// TIA Portal project "FABRICA DE TAPAS - TRANSPORTE -TUNEL DE ENFRIAMIENTO" (V17) (continued)
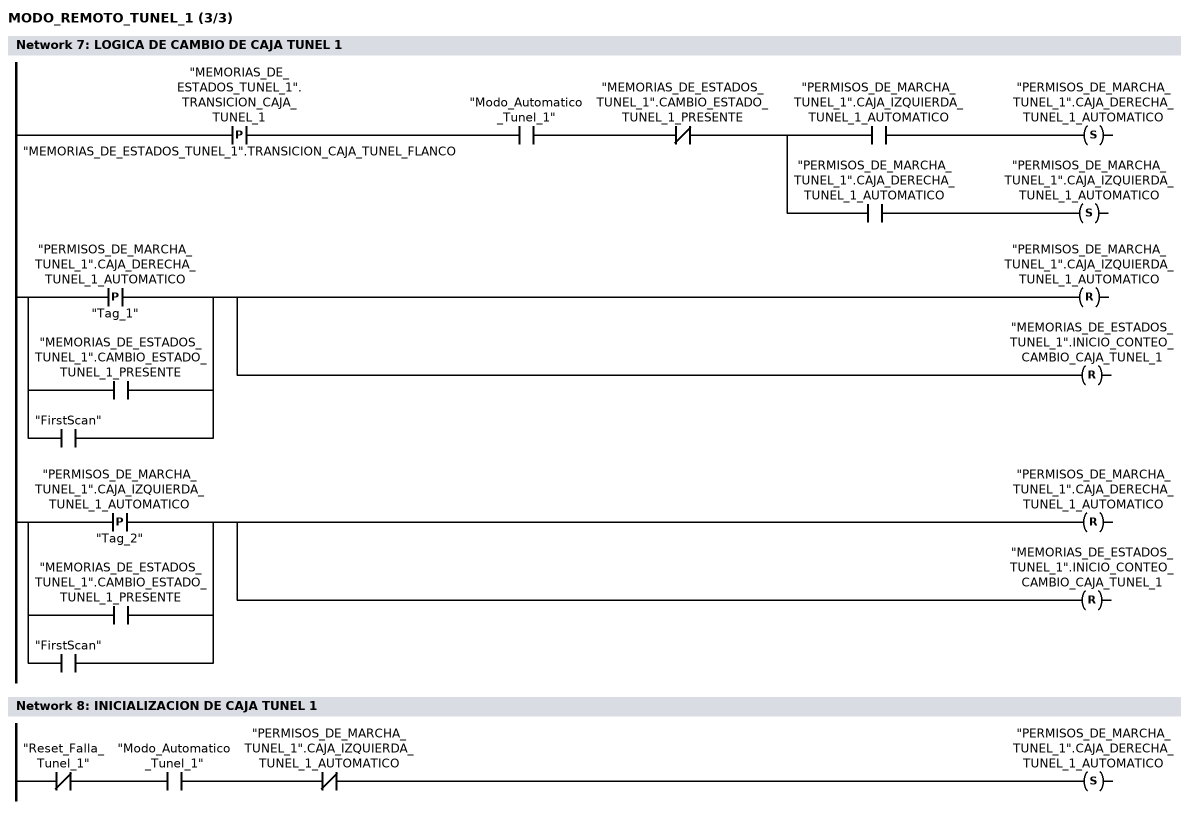
   RUNG wire#powerrail
      P_Contact(operand := "MEMORIAS_DE_ESTADOS_TUNEL_1".TRANSICION_CAJA_TUNEL_1, bit := "MEMORIAS_DE_ESTADOS_TUNEL_1".TRANSICION_CAJA_TUNEL_FLANCO)
      Contact( "Modo_Automatico_Tunel_1" )
      I_Contact( "MEMORIAS_DE_ESTADOS_TUNEL_1".CAMBIO_ESTADO_TUNEL_1_PRESENTE )
      wire#w1
      Contact( "PERMISOS_DE_MARCHA_TUNEL_1".CAJA_IZQUIERDA_TUNEL_1_AUTOMATICO )
      S_Coil( "PERMISOS_DE_MARCHA_TUNEL_1".CAJA_DERECHA_TUNEL_1_AUTOMATICO )
   END_RUNG
   RUNG wire#w1
      Contact( "PERMISOS_DE_MARCHA_TUNEL_1".CAJA_DERECHA_TUNEL_1_AUTOMATICO )
      S_Coil( "PERMISOS_DE_MARCHA_TUNEL_1".CAJA_IZQUIERDA_TUNEL_1_AUTOMATICO )
   END_RUNG
   RUNG wire#powerrail
      P_Contact(operand := "PERMISOS_DE_MARCHA_TUNEL_1".CAJA_DERECHA_TUNEL_1_AUTOMATICO, bit := "Tag_1")
      wire#w2
      R_Coil( "PERMISOS_DE_MARCHA_TUNEL_1".CAJA_IZQUIERDA_TUNEL_1_AUTOMATICO )
   END_RUNG
   RUNG wire#powerrail
      Contact( "MEMORIAS_DE_ESTADOS_TUNEL_1".CAMBIO_ESTADO_TUNEL_1_PRESENTE )
   END_RUNG wire#w2
   RUNG wire#powerrail
      Contact( "FirstScan" )
   END_RUNG wire#w2
   RUNG wire#w2
      R_Coil( "MEMORIAS_DE_ESTADOS_TUNEL_1".INICIO_CONTEO_CAMBIO_CAJA_TUNEL_1 )
   END_RUNG
   RUNG wire#powerrail
      P_Contact(operand := "PERMISOS_DE_MARCHA_TUNEL_1".CAJA_IZQUIERDA_TUNEL_1_AUTOMATICO, bit := "Tag_2")
      wire#w3
      R_Coil( "PERMISOS_DE_MARCHA_TUNEL_1".CAJA_DERECHA_TUNEL_1_AUTOMATICO )
   END_RUNG
   RUNG wire#powerrail
      Contact( "MEMORIAS_DE_ESTADOS_TUNEL_1".CAMBIO_ESTADO_TUNEL_1_PRESENTE )
   END_RUNG wire#w3
   RUNG wire#powerrail
      Contact( "FirstScan" )
   END_RUNG wire#w3
   RUNG wire#w3
      R_Coil( "MEMORIAS_DE_ESTADOS_TUNEL_1".INICIO_CONTEO_CAMBIO_CAJA_TUNEL_1 )
   END_RUNG
   // the same network as SCL:
   #_w1 := "MEMORIAS_DE_ESTADOS_TUNEL_1".TRANSICION_CAJA_TUNEL_1 AND NOT "MEMORIAS_DE_ESTADOS_TUNEL_1".TRANSICION_CAJA_TUNEL_FLANCO;   // rising edge of "MEMORIAS_DE_ESTADOS_TUNEL_1".TRANSICION_CAJA_TUNEL_1
   "MEMORIAS_DE_ESTADOS_TUNEL_1".TRANSICION_CAJA_TUNEL_FLANCO := "MEMORIAS_DE_ESTADOS_TUNEL_1".TRANSICION_CAJA_TUNEL_1;
   #_w2 := #_w1 AND "Modo_Automatico_Tunel_1" AND NOT "MEMORIAS_DE_ESTADOS_TUNEL_1".CAMBIO_ESTADO_TUNEL_1_PRESENTE;
   IF #_w2 AND "PERMISOS_DE_MARCHA_TUNEL_1".CAJA_IZQUIERDA_TUNEL_1_AUTOMATICO THEN
       "PERMISOS_DE_MARCHA_TUNEL_1".CAJA_DERECHA_TUNEL_1_AUTOMATICO := TRUE;
   END_IF;
   IF #_w2 AND "PERMISOS_DE_MARCHA_TUNEL_1".CAJA_DERECHA_TUNEL_1_AUTOMATICO THEN
       "PERMISOS_DE_MARCHA_TUNEL_1".CAJA_IZQUIERDA_TUNEL_1_AUTOMATICO := TRUE;
   END_IF;
   #_w3 := "PERMISOS_DE_MARCHA_TUNEL_1".CAJA_DERECHA_TUNEL_1_AUTOMATICO AND NOT "Tag_1";   // rising edge of "PERMISOS_DE_MARCHA_TUNEL_1".CAJA_DERECHA_TUNEL_1_AUTOMATICO
   "Tag_1" := "PERMISOS_DE_MARCHA_TUNEL_1".CAJA_DERECHA_TUNEL_1_AUTOMATICO;
   IF #_w3 OR "MEMORIAS_DE_ESTADOS_TUNEL_1".CAMBIO_ESTADO_TUNEL_1_PRESENTE OR "FirstScan" THEN
       "PERMISOS_DE_MARCHA_TUNEL_1".CAJA_IZQUIERDA_TUNEL_1_AUTOMATICO := FALSE;
       "MEMORIAS_DE_ESTADOS_TUNEL_1".INICIO_CONTEO_CAMBIO_CAJA_TUNEL_1 := FALSE;
   END_IF;
   #_w4 := "PERMISOS_DE_MARCHA_TUNEL_1".CAJA_IZQUIERDA_TUNEL_1_AUTOMATICO AND NOT "Tag_2";   // rising edge of "PERMISOS_DE_MARCHA_TUNEL_1".CAJA_IZQUIERDA_TUNEL_1_AUTOMATICO
   "Tag_2" := "PERMISOS_DE_MARCHA_TUNEL_1".CAJA_IZQUIERDA_TUNEL_1_AUTOMATICO;
   IF #_w4 OR "MEMORIAS_DE_ESTADOS_TUNEL_1".CAMBIO_ESTADO_TUNEL_1_PRESENTE OR "FirstScan" THEN
       "PERMISOS_DE_MARCHA_TUNEL_1".CAJA_DERECHA_TUNEL_1_AUTOMATICO := FALSE;
       "MEMORIAS_DE_ESTADOS_TUNEL_1".INICIO_CONTEO_CAMBIO_CAJA_TUNEL_1 := FALSE;
   END_IF;
END_REGION

REGION Network 8: INICIALIZACION DE CAJA TUNEL 1
   RUNG wire#powerrail
      I_Contact( "Reset_Falla_Tunel_1" )
      Contact( "Modo_Automatico_Tunel_1" )
      I_Contact( "PERMISOS_DE_MARCHA_TUNEL_1".CAJA_IZQUIERDA_TUNEL_1_AUTOMATICO )
      S_Coil( "PERMISOS_DE_MARCHA_TUNEL_1".CAJA_DERECHA_TUNEL_1_AUTOMATICO )
   END_RUNG
   // the same network as SCL:
   IF NOT "Reset_Falla_Tunel_1" AND "Modo_Automatico_Tunel_1" AND NOT "PERMISOS_DE_MARCHA_TUNEL_1".CAJA_IZQUIERDA_TUNEL_1_AUTOMATICO THEN
       "PERMISOS_DE_MARCHA_TUNEL_1".CAJA_DERECHA_TUNEL_1_AUTOMATICO := TRUE;
   END_IF;
END_REGION
END_FUNCTION

FUNCTION "MODO_REMOTO_TUNEL_2" : Void   // FC2, LAD
{ S7_Optimized_Access := 'TRUE' }
VERSION : 0.1
   VAR_TEMP   // added for the SCL form of the ladder/FBD networks
      _w1 : Bool;
      _w2 : Bool;
      _w3 : Bool;
      _w4 : Bool;
   END_VAR
BEGIN

REGION Network 1
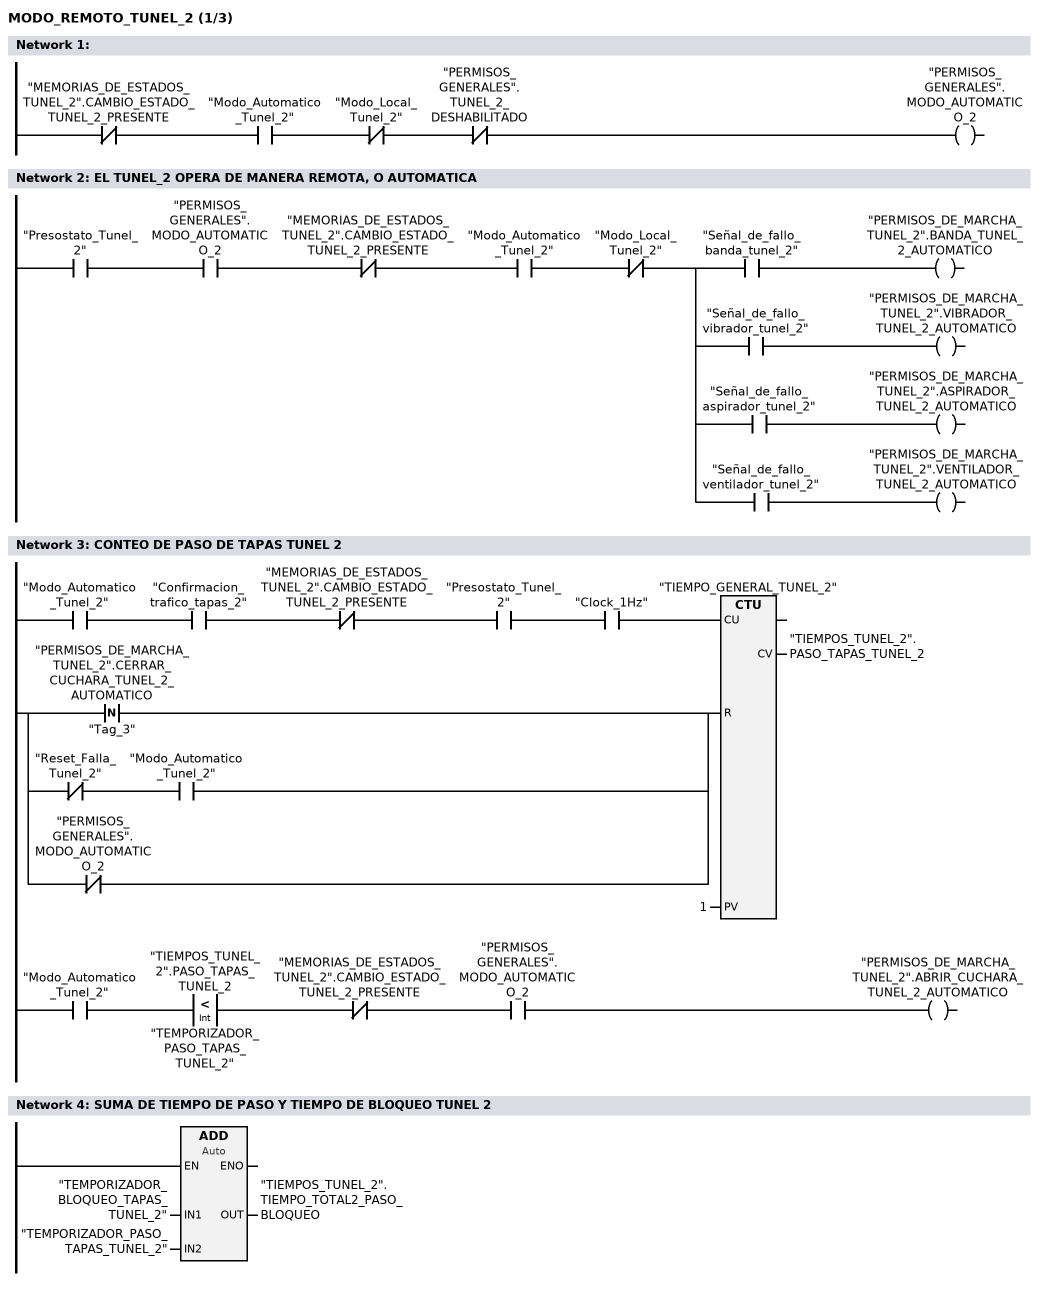
   RUNG wire#powerrail
      I_Contact( "MEMORIAS_DE_ESTADOS_TUNEL_2".CAMBIO_ESTADO_TUNEL_2_PRESENTE )
      Contact( "Modo_Automatico_Tunel_2" )
      I_Contact( "Modo_Local_Tunel_2" )
      I_Contact( "PERMISOS_GENERALES".TUNEL_2_DESHABILITADO )
      Coil( "PERMISOS_GENERALES".MODO_AUTOMATICO_2 )
   END_RUNG
   // the same network as SCL:
   "PERMISOS_GENERALES".MODO_AUTOMATICO_2 := NOT "MEMORIAS_DE_ESTADOS_TUNEL_2".CAMBIO_ESTADO_TUNEL_2_PRESENTE AND "Modo_Automatico_Tunel_2" AND NOT "Modo_Local_Tunel_2" AND NOT "PERMISOS_GENERALES".TUNEL_2_DESHABILITADO;
END_REGION

REGION Network 2: EL TUNEL_2 OPERA DE MANERA REMOTA, O AUTOMATICA
   RUNG wire#powerrail
      Contact( "Presostato_Tunel_2" )
      Contact( "PERMISOS_GENERALES".MODO_AUTOMATICO_2 )
      I_Contact( "MEMORIAS_DE_ESTADOS_TUNEL_2".CAMBIO_ESTADO_TUNEL_2_PRESENTE )
      Contact( "Modo_Automatico_Tunel_2" )
      I_Contact( "Modo_Local_Tunel_2" )
      wire#w1
      Contact( "Señal_de_fallo_banda_tunel_2" )
      Coil( "PERMISOS_DE_MARCHA_TUNEL_2".BANDA_TUNEL_2_AUTOMATICO )
   END_RUNG
   RUNG wire#w1
      Contact( "Señal_de_fallo_vibrador_tunel_2" )
      Coil( "PERMISOS_DE_MARCHA_TUNEL_2".VIBRADOR_TUNEL_2_AUTOMATICO )
   END_RUNG
   RUNG wire#w1
      Contact( "Señal_de_fallo_aspirador_tunel_2" )
      Coil( "PERMISOS_DE_MARCHA_TUNEL_2".ASPIRADOR_TUNEL_2_AUTOMATICO )
   END_RUNG
   RUNG wire#w1
      Contact( "Señal_de_fallo_ventilador_tunel_2" )
      Coil( "PERMISOS_DE_MARCHA_TUNEL_2".VENTILADOR_TUNEL_2_AUTOMATICO )
   END_RUNG
   // the same network as SCL:
   #_w1 := "Presostato_Tunel_2" AND "PERMISOS_GENERALES".MODO_AUTOMATICO_2 AND NOT "MEMORIAS_DE_ESTADOS_TUNEL_2".CAMBIO_ESTADO_TUNEL_2_PRESENTE AND "Modo_Automatico_Tunel_2" AND NOT "Modo_Local_Tunel_2";
   "PERMISOS_DE_MARCHA_TUNEL_2".BANDA_TUNEL_2_AUTOMATICO := #_w1 AND "Señal_de_fallo_banda_tunel_2";
   "PERMISOS_DE_MARCHA_TUNEL_2".VIBRADOR_TUNEL_2_AUTOMATICO := #_w1 AND "Señal_de_fallo_vibrador_tunel_2";
   "PERMISOS_DE_MARCHA_TUNEL_2".ASPIRADOR_TUNEL_2_AUTOMATICO := #_w1 AND "Señal_de_fallo_aspirador_tunel_2";
   "PERMISOS_DE_MARCHA_TUNEL_2".VENTILADOR_TUNEL_2_AUTOMATICO := #_w1 AND "Señal_de_fallo_ventilador_tunel_2";
END_REGION

REGION Network 3: CONTEO DE PASO DE TAPAS TUNEL 2
   #_w1 := NOT "PERMISOS_DE_MARCHA_TUNEL_2".CERRAR_CUCHARA_TUNEL_2_AUTOMATICO AND "Tag_3";   // falling edge of "PERMISOS_DE_MARCHA_TUNEL_2".CERRAR_CUCHARA_TUNEL_2_AUTOMATICO
   "Tag_3" := "PERMISOS_DE_MARCHA_TUNEL_2".CERRAR_CUCHARA_TUNEL_2_AUTOMATICO;
   "TIEMPO_GENERAL_TUNEL_2".CTU(CU := "Modo_Automatico_Tunel_2" AND "Confirmacion_trafico_tapas_2" AND NOT "MEMORIAS_DE_ESTADOS_TUNEL_2".CAMBIO_ESTADO_TUNEL_2_PRESENTE AND "Presostato_Tunel_2" AND "Clock_1Hz",
                           R := #_w1 OR (NOT "Reset_Falla_Tunel_2" AND "Modo_Automatico_Tunel_2") OR NOT "PERMISOS_GENERALES".MODO_AUTOMATICO_2,
                           PV := 1,
                           CV => "TIEMPOS_TUNEL_2".PASO_TAPAS_TUNEL_2);
   "PERMISOS_DE_MARCHA_TUNEL_2".ABRIR_CUCHARA_TUNEL_2_AUTOMATICO := "Modo_Automatico_Tunel_2" AND ("TIEMPOS_TUNEL_2".PASO_TAPAS_TUNEL_2 < "TEMPORIZADOR_PASO_TAPAS_TUNEL_2") AND NOT "MEMORIAS_DE_ESTADOS_TUNEL_2".CAMBIO_ESTADO_TUNEL_2_PRESENTE AND "PERMISOS_GENERALES".MODO_AUTOMATICO_2;
END_REGION

REGION Network 4: SUMA DE TIEMPO DE PASO Y TIEMPO DE BLOQUEO TUNEL 2
   RUNG wire#powerrail
      Add(in1 := "TEMPORIZADOR_BLOQUEO_TAPAS_TUNEL_2", in2 := "TEMPORIZADOR_PASO_TAPAS_TUNEL_2", out => "TIEMPOS_TUNEL_2".TIEMPO_TOTAL2_PASO_BLOQUEO)
   END_RUNG
   // the same network as SCL:
   "TIEMPOS_TUNEL_2".TIEMPO_TOTAL2_PASO_BLOQUEO := "TEMPORIZADOR_BLOQUEO_TAPAS_TUNEL_2" + "TEMPORIZADOR_PASO_TAPAS_TUNEL_2";
END_REGION

REGION Network 5: CIERRE DE CUCHARRA PARA BLOQUEO DE TAPAS TUNEL 2
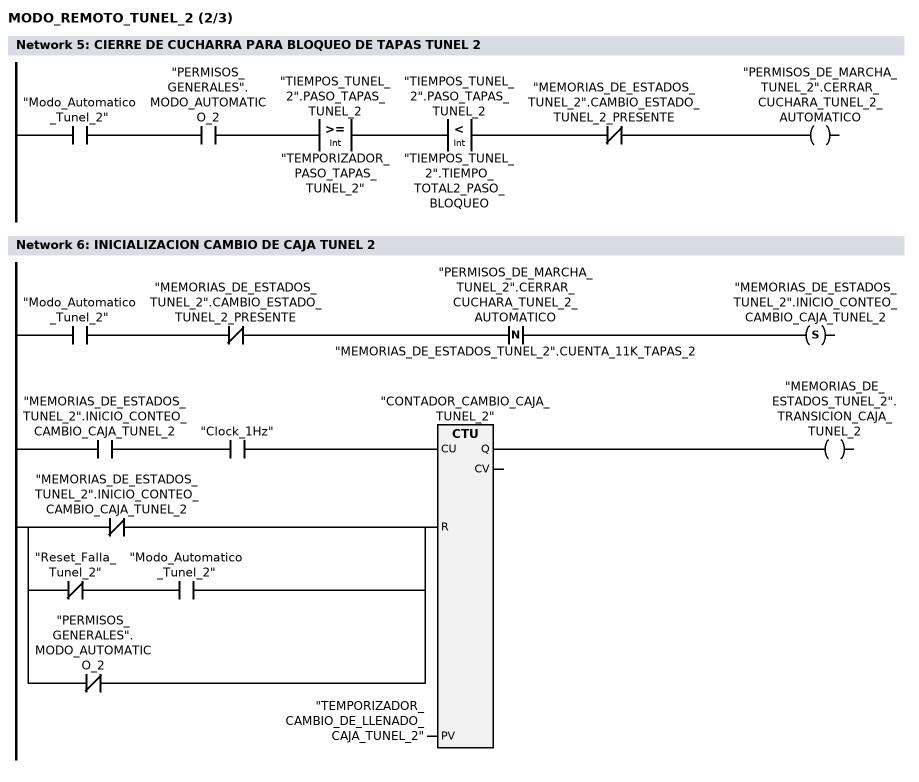
   RUNG wire#powerrail
      Contact( "Modo_Automatico_Tunel_2" )
      Contact( "PERMISOS_GENERALES".MODO_AUTOMATICO_2 )
      { S7_Templates := "SrcType := Int" } GE_Contact(in1 := "TIEMPOS_TUNEL_2".PASO_TAPAS_TUNEL_2, in2 := "TEMPORIZADOR_PASO_TAPAS_TUNEL_2")
      { S7_Templates := "SrcType := Int" } LT_Contact(in1 := "TIEMPOS_TUNEL_2".PASO_TAPAS_TUNEL_2, in2 := "TIEMPOS_TUNEL_2".TIEMPO_TOTAL2_PASO_BLOQUEO)
      I_Contact( "MEMORIAS_DE_ESTADOS_TUNEL_2".CAMBIO_ESTADO_TUNEL_2_PRESENTE )
      Coil( "PERMISOS_DE_MARCHA_TUNEL_2".CERRAR_CUCHARA_TUNEL_2_AUTOMATICO )
   END_RUNG
   // the same network as SCL:
   "PERMISOS_DE_MARCHA_TUNEL_2".CERRAR_CUCHARA_TUNEL_2_AUTOMATICO := "Modo_Automatico_Tunel_2" AND "PERMISOS_GENERALES".MODO_AUTOMATICO_2 AND ("TIEMPOS_TUNEL_2".PASO_TAPAS_TUNEL_2 >= "TEMPORIZADOR_PASO_TAPAS_TUNEL_2") AND ("TIEMPOS_TUNEL_2".PASO_TAPAS_TUNEL_2 < "TIEMPOS_TUNEL_2".TIEMPO_TOTAL2_PASO_BLOQUEO) AND NOT "MEMORIAS_DE_ESTADOS_TUNEL_2".CAMBIO_ESTADO_TUNEL_2_PRESENTE;
END_REGION

REGION Network 6: INICIALIZACION CAMBIO DE CAJA TUNEL 2
   #_w1 := "Modo_Automatico_Tunel_2" AND NOT "MEMORIAS_DE_ESTADOS_TUNEL_2".CAMBIO_ESTADO_TUNEL_2_PRESENTE AND NOT "PERMISOS_DE_MARCHA_TUNEL_2".CERRAR_CUCHARA_TUNEL_2_AUTOMATICO AND "MEMORIAS_DE_ESTADOS_TUNEL_2".CUENTA_11K_TAPAS_2;   // falling edge of "PERMISOS_DE_MARCHA_TUNEL_2".CERRAR_CUCHARA_TUNEL_2_AUTOMATICO
   "MEMORIAS_DE_ESTADOS_TUNEL_2".CUENTA_11K_TAPAS_2 := "PERMISOS_DE_MARCHA_TUNEL_2".CERRAR_CUCHARA_TUNEL_2_AUTOMATICO;
   IF #_w1 THEN "MEMORIAS_DE_ESTADOS_TUNEL_2".INICIO_CONTEO_CAMBIO_CAJA_TUNEL_2 := TRUE; END_IF;
   "CONTADOR_CAMBIO_CAJA_TUNEL_2".CTU(CU := "MEMORIAS_DE_ESTADOS_TUNEL_2".INICIO_CONTEO_CAMBIO_CAJA_TUNEL_2 AND "Clock_1Hz",
                           R := NOT "MEMORIAS_DE_ESTADOS_TUNEL_2".INICIO_CONTEO_CAMBIO_CAJA_TUNEL_2 OR (NOT "Reset_Falla_Tunel_2" AND "Modo_Automatico_Tunel_2") OR NOT "PERMISOS_GENERALES".MODO_AUTOMATICO_2,
                           PV := "TEMPORIZADOR_CAMBIO_DE_LLENADO_CAJA_TUNEL_2");
   "MEMORIAS_DE_ESTADOS_TUNEL_2".TRANSICION_CAJA_TUNEL_2 := "CONTADOR_CAMBIO_CAJA_TUNEL_2".Q;
END_REGION

REGION Network 7: LOGICA DE CAMBIO DE CAJA TUNEL 2
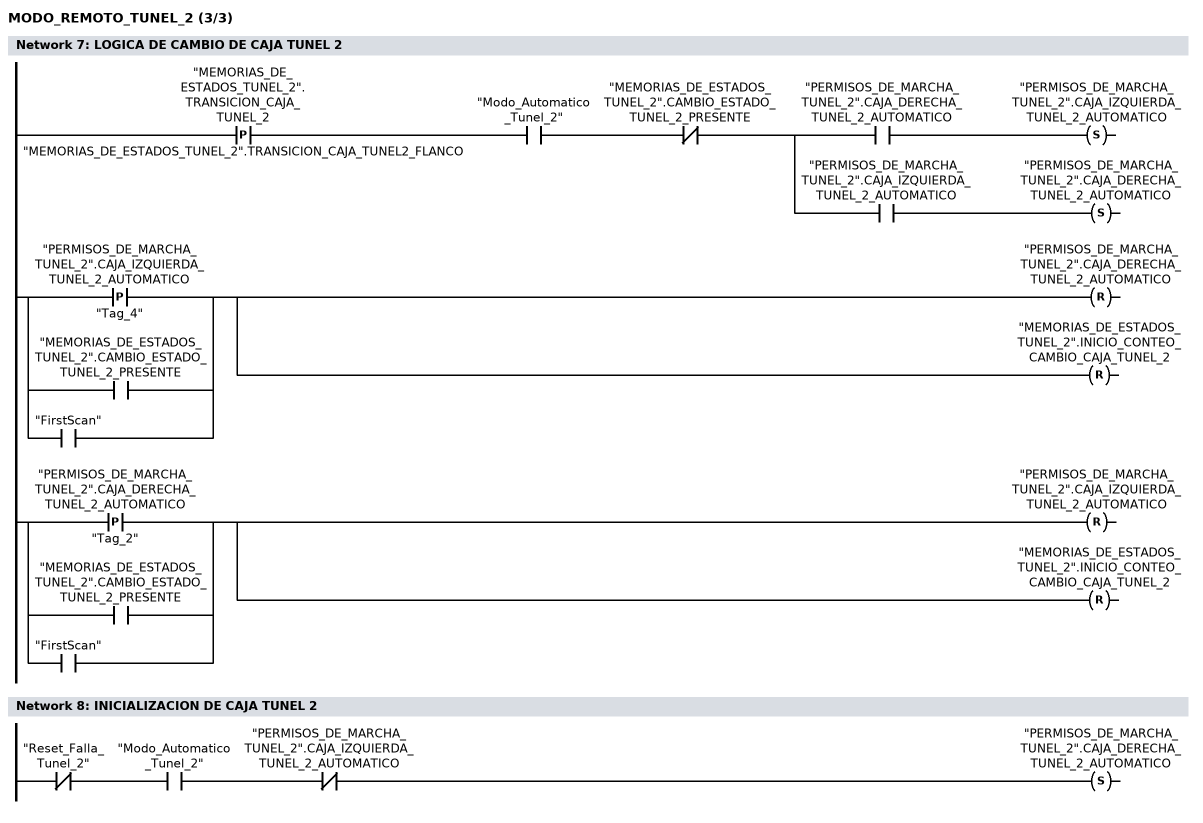
   RUNG wire#powerrail
      P_Contact(operand := "MEMORIAS_DE_ESTADOS_TUNEL_2".TRANSICION_CAJA_TUNEL_2, bit := "MEMORIAS_DE_ESTADOS_TUNEL_2".TRANSICION_CAJA_TUNEL2_FLANCO)
      Contact( "Modo_Automatico_Tunel_2" )
      I_Contact( "MEMORIAS_DE_ESTADOS_TUNEL_2".CAMBIO_ESTADO_TUNEL_2_PRESENTE )
      wire#w1
      Contact( "PERMISOS_DE_MARCHA_TUNEL_2".CAJA_DERECHA_TUNEL_2_AUTOMATICO )
      S_Coil( "PERMISOS_DE_MARCHA_TUNEL_2".CAJA_IZQUIERDA_TUNEL_2_AUTOMATICO )
   END_RUNG
   RUNG wire#w1
      Contact( "PERMISOS_DE_MARCHA_TUNEL_2".CAJA_IZQUIERDA_TUNEL_2_AUTOMATICO )
      S_Coil( "PERMISOS_DE_MARCHA_TUNEL_2".CAJA_DERECHA_TUNEL_2_AUTOMATICO )
   END_RUNG
   RUNG wire#powerrail
      P_Contact(operand := "PERMISOS_DE_MARCHA_TUNEL_2".CAJA_IZQUIERDA_TUNEL_2_AUTOMATICO, bit := "Tag_4")
      wire#w2
      R_Coil( "PERMISOS_DE_MARCHA_TUNEL_2".CAJA_DERECHA_TUNEL_2_AUTOMATICO )
   END_RUNG
   RUNG wire#powerrail
      Contact( "MEMORIAS_DE_ESTADOS_TUNEL_2".CAMBIO_ESTADO_TUNEL_2_PRESENTE )
   END_RUNG wire#w2
   RUNG wire#powerrail
      Contact( "FirstScan" )
   END_RUNG wire#w2
   RUNG wire#w2
      R_Coil( "MEMORIAS_DE_ESTADOS_TUNEL_2".INICIO_CONTEO_CAMBIO_CAJA_TUNEL_2 )
   END_RUNG
   RUNG wire#powerrail
      P_Contact(operand := "PERMISOS_DE_MARCHA_TUNEL_2".CAJA_DERECHA_TUNEL_2_AUTOMATICO, bit := "Tag_2")
      wire#w3
      R_Coil( "PERMISOS_DE_MARCHA_TUNEL_2".CAJA_IZQUIERDA_TUNEL_2_AUTOMATICO )
   END_RUNG
   RUNG wire#powerrail
      Contact( "MEMORIAS_DE_ESTADOS_TUNEL_2".CAMBIO_ESTADO_TUNEL_2_PRESENTE )
   END_RUNG wire#w3
   RUNG wire#powerrail
      Contact( "FirstScan" )
   END_RUNG wire#w3
   RUNG wire#w3
      R_Coil( "MEMORIAS_DE_ESTADOS_TUNEL_2".INICIO_CONTEO_CAMBIO_CAJA_TUNEL_2 )
   END_RUNG
   // the same network as SCL:
   #_w1 := "MEMORIAS_DE_ESTADOS_TUNEL_2".TRANSICION_CAJA_TUNEL_2 AND NOT "MEMORIAS_DE_ESTADOS_TUNEL_2".TRANSICION_CAJA_TUNEL2_FLANCO;   // rising edge of "MEMORIAS_DE_ESTADOS_TUNEL_2".TRANSICION_CAJA_TUNEL_2
   "MEMORIAS_DE_ESTADOS_TUNEL_2".TRANSICION_CAJA_TUNEL2_FLANCO := "MEMORIAS_DE_ESTADOS_TUNEL_2".TRANSICION_CAJA_TUNEL_2;
   #_w2 := #_w1 AND "Modo_Automatico_Tunel_2" AND NOT "MEMORIAS_DE_ESTADOS_TUNEL_2".CAMBIO_ESTADO_TUNEL_2_PRESENTE;
   IF #_w2 AND "PERMISOS_DE_MARCHA_TUNEL_2".CAJA_DERECHA_TUNEL_2_AUTOMATICO THEN
       "PERMISOS_DE_MARCHA_TUNEL_2".CAJA_IZQUIERDA_TUNEL_2_AUTOMATICO := TRUE;
   END_IF;
   IF #_w2 AND "PERMISOS_DE_MARCHA_TUNEL_2".CAJA_IZQUIERDA_TUNEL_2_AUTOMATICO THEN
       "PERMISOS_DE_MARCHA_TUNEL_2".CAJA_DERECHA_TUNEL_2_AUTOMATICO := TRUE;
   END_IF;
   #_w3 := "PERMISOS_DE_MARCHA_TUNEL_2".CAJA_IZQUIERDA_TUNEL_2_AUTOMATICO AND NOT "Tag_4";   // rising edge of "PERMISOS_DE_MARCHA_TUNEL_2".CAJA_IZQUIERDA_TUNEL_2_AUTOMATICO
   "Tag_4" := "PERMISOS_DE_MARCHA_TUNEL_2".CAJA_IZQUIERDA_TUNEL_2_AUTOMATICO;
   IF #_w3 OR "MEMORIAS_DE_ESTADOS_TUNEL_2".CAMBIO_ESTADO_TUNEL_2_PRESENTE OR "FirstScan" THEN
       "PERMISOS_DE_MARCHA_TUNEL_2".CAJA_DERECHA_TUNEL_2_AUTOMATICO := FALSE;
       "MEMORIAS_DE_ESTADOS_TUNEL_2".INICIO_CONTEO_CAMBIO_CAJA_TUNEL_2 := FALSE;
   END_IF;
   #_w4 := "PERMISOS_DE_MARCHA_TUNEL_2".CAJA_DERECHA_TUNEL_2_AUTOMATICO AND NOT "Tag_2";   // rising edge of "PERMISOS_DE_MARCHA_TUNEL_2".CAJA_DERECHA_TUNEL_2_AUTOMATICO
   "Tag_2" := "PERMISOS_DE_MARCHA_TUNEL_2".CAJA_DERECHA_TUNEL_2_AUTOMATICO;
   IF #_w4 OR "MEMORIAS_DE_ESTADOS_TUNEL_2".CAMBIO_ESTADO_TUNEL_2_PRESENTE OR "FirstScan" THEN
       "PERMISOS_DE_MARCHA_TUNEL_2".CAJA_IZQUIERDA_TUNEL_2_AUTOMATICO := FALSE;
       "MEMORIAS_DE_ESTADOS_TUNEL_2".INICIO_CONTEO_CAMBIO_CAJA_TUNEL_2 := FALSE;
   END_IF;
END_REGION

REGION Network 8: INICIALIZACION DE CAJA TUNEL 2
   RUNG wire#powerrail
      I_Contact( "Reset_Falla_Tunel_2" )
      Contact( "Modo_Automatico_Tunel_2" )
      I_Contact( "PERMISOS_DE_MARCHA_TUNEL_2".CAJA_IZQUIERDA_TUNEL_2_AUTOMATICO )
      S_Coil( "PERMISOS_DE_MARCHA_TUNEL_2".CAJA_DERECHA_TUNEL_2_AUTOMATICO )
   END_RUNG
   // the same network as SCL:
   IF NOT "Reset_Falla_Tunel_2" AND "Modo_Automatico_Tunel_2" AND NOT "PERMISOS_DE_MARCHA_TUNEL_2".CAJA_IZQUIERDA_TUNEL_2_AUTOMATICO THEN
       "PERMISOS_DE_MARCHA_TUNEL_2".CAJA_DERECHA_TUNEL_2_AUTOMATICO := TRUE;
   END_IF;
END_REGION
END_FUNCTION

FUNCTION "OPERACION_MODO_LOCAL_TUNEL_1" : Void   // FC3, LAD
{ S7_Optimized_Access := 'TRUE' }
VERSION : 0.1
BEGIN

REGION Network 1
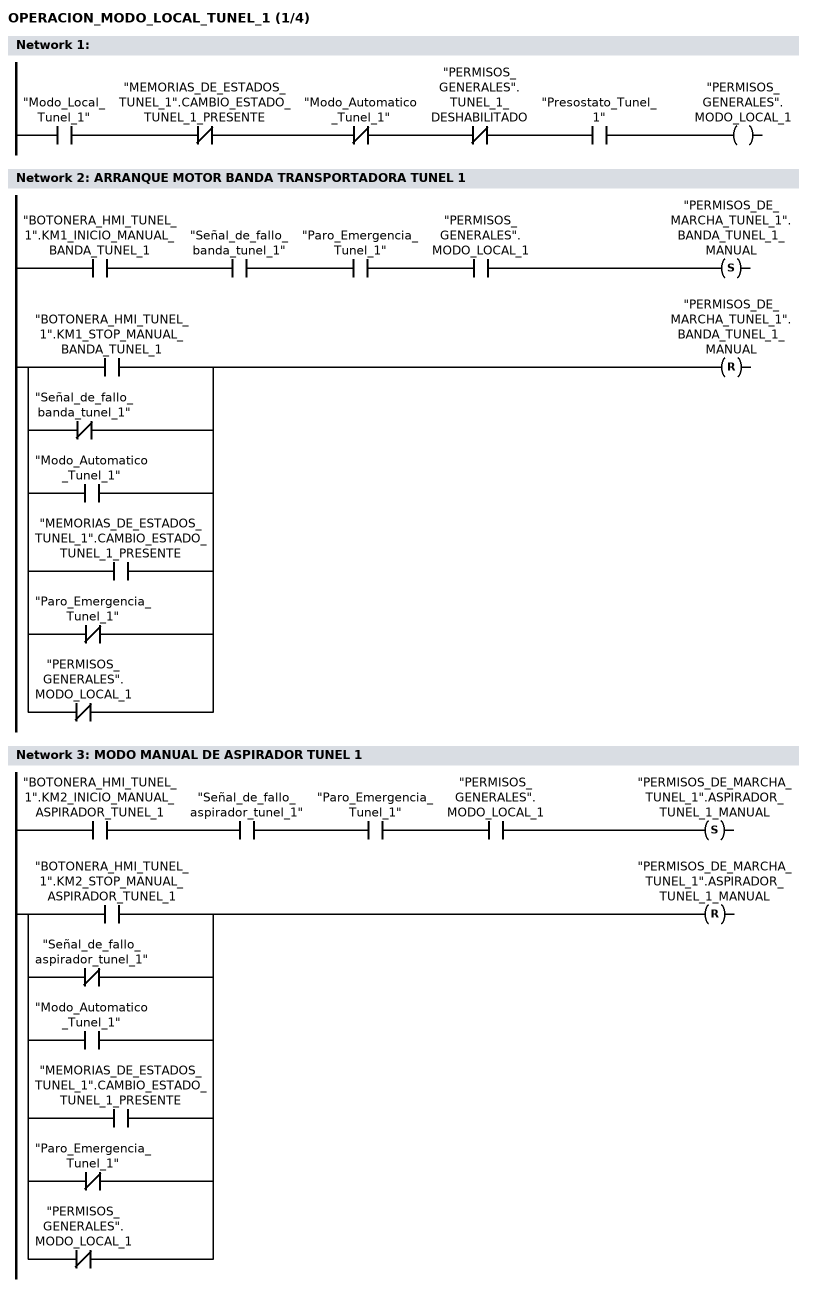
   RUNG wire#powerrail
      Contact( "Modo_Local_Tunel_1" )
      I_Contact( "MEMORIAS_DE_ESTADOS_TUNEL_1".CAMBIO_ESTADO_TUNEL_1_PRESENTE )
      I_Contact( "Modo_Automatico_Tunel_1" )
      I_Contact( "PERMISOS_GENERALES".TUNEL_1_DESHABILITADO )
      Contact( "Presostato_Tunel_1" )
      Coil( "PERMISOS_GENERALES".MODO_LOCAL_1 )
   END_RUNG
   // the same network as SCL:
   "PERMISOS_GENERALES".MODO_LOCAL_1 := "Modo_Local_Tunel_1" AND NOT "MEMORIAS_DE_ESTADOS_TUNEL_1".CAMBIO_ESTADO_TUNEL_1_PRESENTE AND NOT "Modo_Automatico_Tunel_1" AND NOT "PERMISOS_GENERALES".TUNEL_1_DESHABILITADO AND "Presostato_Tunel_1";
END_REGION

REGION Network 2: ARRANQUE MOTOR BANDA TRANSPORTADORA TUNEL 1
   RUNG wire#powerrail
      Contact( "BOTONERA_HMI_TUNEL_1".KM1_INICIO_MANUAL_BANDA_TUNEL_1 )
      Contact( "Señal_de_fallo_banda_tunel_1" )
      Contact( "Paro_Emergencia_Tunel_1" )
      Contact( "PERMISOS_GENERALES".MODO_LOCAL_1 )
      S_Coil( "PERMISOS_DE_MARCHA_TUNEL_1".BANDA_TUNEL_1_MANUAL )
   END_RUNG
   RUNG wire#powerrail
      Contact( "BOTONERA_HMI_TUNEL_1".KM1_STOP_MANUAL_BANDA_TUNEL_1 )
      wire#w1
      R_Coil( "PERMISOS_DE_MARCHA_TUNEL_1".BANDA_TUNEL_1_MANUAL )
   END_RUNG
   RUNG wire#powerrail
      I_Contact( "Señal_de_fallo_banda_tunel_1" )
   END_RUNG wire#w1
   RUNG wire#powerrail
      Contact( "Modo_Automatico_Tunel_1" )
   END_RUNG wire#w1
   RUNG wire#powerrail
      Contact( "MEMORIAS_DE_ESTADOS_TUNEL_1".CAMBIO_ESTADO_TUNEL_1_PRESENTE )
   END_RUNG wire#w1
   RUNG wire#powerrail
      I_Contact( "Paro_Emergencia_Tunel_1" )
   END_RUNG wire#w1
   RUNG wire#powerrail
      I_Contact( "PERMISOS_GENERALES".MODO_LOCAL_1 )
   END_RUNG wire#w1
   // the same network as SCL:
   IF "BOTONERA_HMI_TUNEL_1".KM1_INICIO_MANUAL_BANDA_TUNEL_1 AND "Señal_de_fallo_banda_tunel_1" AND "Paro_Emergencia_Tunel_1" AND "PERMISOS_GENERALES".MODO_LOCAL_1 THEN
       "PERMISOS_DE_MARCHA_TUNEL_1".BANDA_TUNEL_1_MANUAL := TRUE;
   END_IF;
   IF "BOTONERA_HMI_TUNEL_1".KM1_STOP_MANUAL_BANDA_TUNEL_1 OR NOT "Señal_de_fallo_banda_tunel_1" OR "Modo_Automatico_Tunel_1" OR "MEMORIAS_DE_ESTADOS_TUNEL_1".CAMBIO_ESTADO_TUNEL_1_PRESENTE OR NOT "Paro_Emergencia_Tunel_1" OR NOT "PERMISOS_GENERALES".MODO_LOCAL_1 THEN
       "PERMISOS_DE_MARCHA_TUNEL_1".BANDA_TUNEL_1_MANUAL := FALSE;
   END_IF;
END_REGION

REGION Network 3: MODO MANUAL DE ASPIRADOR TUNEL 1
   RUNG wire#powerrail
      Contact( "BOTONERA_HMI_TUNEL_1".KM2_INICIO_MANUAL_ASPIRADOR_TUNEL_1 )
      Contact( "Señal_de_fallo_aspirador_tunel_1" )
      Contact( "Paro_Emergencia_Tunel_1" )
      Contact( "PERMISOS_GENERALES".MODO_LOCAL_1 )
      S_Coil( "PERMISOS_DE_MARCHA_TUNEL_1".ASPIRADOR_TUNEL_1_MANUAL )
   END_RUNG
   RUNG wire#powerrail
      Contact( "BOTONERA_HMI_TUNEL_1".KM2_STOP_MANUAL_ASPIRADOR_TUNEL_1 )
      wire#w1
      R_Coil( "PERMISOS_DE_MARCHA_TUNEL_1".ASPIRADOR_TUNEL_1_MANUAL )
   END_RUNG
   RUNG wire#powerrail
      I_Contact( "Señal_de_fallo_aspirador_tunel_1" )
   END_RUNG wire#w1
   RUNG wire#powerrail
      Contact( "Modo_Automatico_Tunel_1" )
   END_RUNG wire#w1
   RUNG wire#powerrail
      Contact( "MEMORIAS_DE_ESTADOS_TUNEL_1".CAMBIO_ESTADO_TUNEL_1_PRESENTE )
   END_RUNG wire#w1
   RUNG wire#powerrail
      I_Contact( "Paro_Emergencia_Tunel_1" )
   END_RUNG wire#w1
   RUNG wire#powerrail
      I_Contact( "PERMISOS_GENERALES".MODO_LOCAL_1 )
   END_RUNG wire#w1
   // the same network as SCL:
   IF "BOTONERA_HMI_TUNEL_1".KM2_INICIO_MANUAL_ASPIRADOR_TUNEL_1 AND "Señal_de_fallo_aspirador_tunel_1" AND "Paro_Emergencia_Tunel_1" AND "PERMISOS_GENERALES".MODO_LOCAL_1 THEN
       "PERMISOS_DE_MARCHA_TUNEL_1".ASPIRADOR_TUNEL_1_MANUAL := TRUE;
   END_IF;
   IF "BOTONERA_HMI_TUNEL_1".KM2_STOP_MANUAL_ASPIRADOR_TUNEL_1 OR NOT "Señal_de_fallo_aspirador_tunel_1" OR "Modo_Automatico_Tunel_1" OR "MEMORIAS_DE_ESTADOS_TUNEL_1".CAMBIO_ESTADO_TUNEL_1_PRESENTE OR NOT "Paro_Emergencia_Tunel_1" OR NOT "PERMISOS_GENERALES".MODO_LOCAL_1 THEN
       "PERMISOS_DE_MARCHA_TUNEL_1".ASPIRADOR_TUNEL_1_MANUAL := FALSE;
   END_IF;
END_REGION

REGION Network 4: MODO MANUAL VENTILADOR TUNEL 1
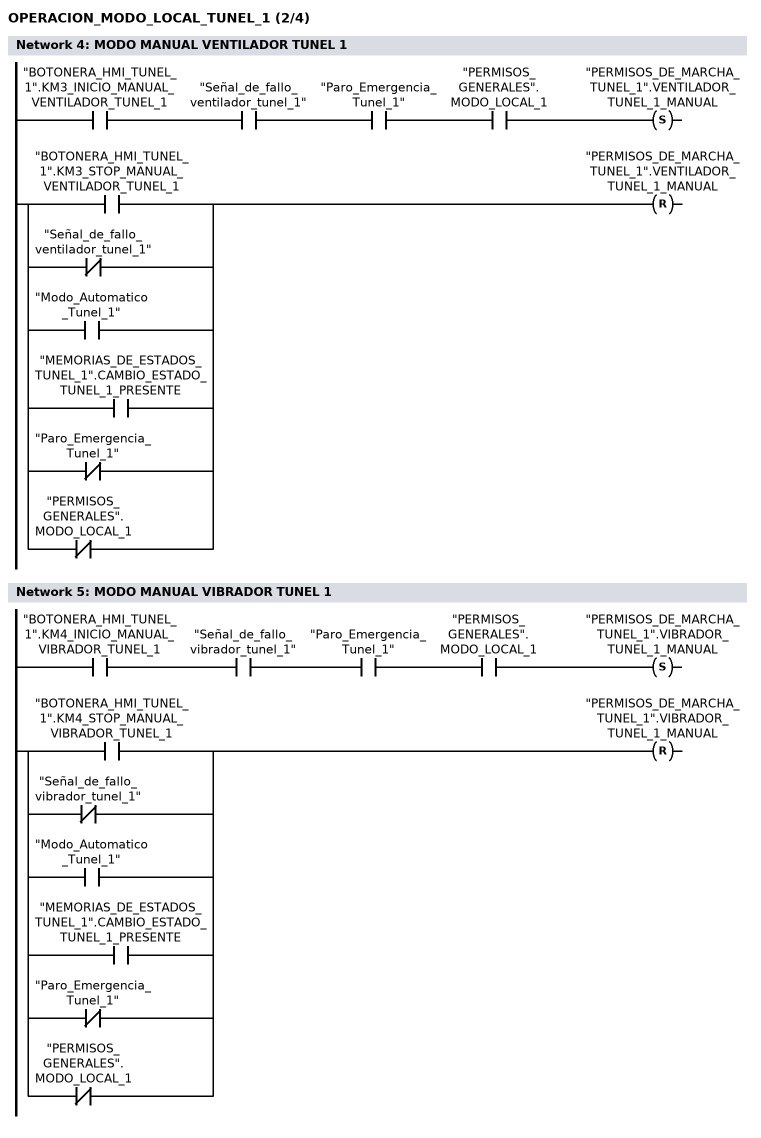
   RUNG wire#powerrail
      Contact( "BOTONERA_HMI_TUNEL_1".KM3_INICIO_MANUAL_VENTILADOR_TUNEL_1 )
      Contact( "Señal_de_fallo_ventilador_tunel_1" )
      Contact( "Paro_Emergencia_Tunel_1" )
      Contact( "PERMISOS_GENERALES".MODO_LOCAL_1 )
      S_Coil( "PERMISOS_DE_MARCHA_TUNEL_1".VENTILADOR_TUNEL_1_MANUAL )
   END_RUNG
   RUNG wire#powerrail
      Contact( "BOTONERA_HMI_TUNEL_1".KM3_STOP_MANUAL_VENTILADOR_TUNEL_1 )
      wire#w1
      R_Coil( "PERMISOS_DE_MARCHA_TUNEL_1".VENTILADOR_TUNEL_1_MANUAL )
   END_RUNG
   RUNG wire#powerrail
      I_Contact( "Señal_de_fallo_ventilador_tunel_1" )
   END_RUNG wire#w1
   RUNG wire#powerrail
      Contact( "Modo_Automatico_Tunel_1" )
   END_RUNG wire#w1
   RUNG wire#powerrail
      Contact( "MEMORIAS_DE_ESTADOS_TUNEL_1".CAMBIO_ESTADO_TUNEL_1_PRESENTE )
   END_RUNG wire#w1
   RUNG wire#powerrail
      I_Contact( "Paro_Emergencia_Tunel_1" )
   END_RUNG wire#w1
   RUNG wire#powerrail
      I_Contact( "PERMISOS_GENERALES".MODO_LOCAL_1 )
   END_RUNG wire#w1
   // the same network as SCL:
   IF "BOTONERA_HMI_TUNEL_1".KM3_INICIO_MANUAL_VENTILADOR_TUNEL_1 AND "Señal_de_fallo_ventilador_tunel_1" AND "Paro_Emergencia_Tunel_1" AND "PERMISOS_GENERALES".MODO_LOCAL_1 THEN
       "PERMISOS_DE_MARCHA_TUNEL_1".VENTILADOR_TUNEL_1_MANUAL := TRUE;
   END_IF;
   IF "BOTONERA_HMI_TUNEL_1".KM3_STOP_MANUAL_VENTILADOR_TUNEL_1 OR NOT "Señal_de_fallo_ventilador_tunel_1" OR "Modo_Automatico_Tunel_1" OR "MEMORIAS_DE_ESTADOS_TUNEL_1".CAMBIO_ESTADO_TUNEL_1_PRESENTE OR NOT "Paro_Emergencia_Tunel_1" OR NOT "PERMISOS_GENERALES".MODO_LOCAL_1 THEN
       "PERMISOS_DE_MARCHA_TUNEL_1".VENTILADOR_TUNEL_1_MANUAL := FALSE;
   END_IF;
END_REGION

REGION Network 5: MODO MANUAL VIBRADOR TUNEL 1
   RUNG wire#powerrail
      Contact( "BOTONERA_HMI_TUNEL_1".KM4_INICIO_MANUAL_VIBRADOR_TUNEL_1 )
      Contact( "Señal_de_fallo_vibrador_tunel_1" )
      Contact( "Paro_Emergencia_Tunel_1" )
      Contact( "PERMISOS_GENERALES".MODO_LOCAL_1 )
      S_Coil( "PERMISOS_DE_MARCHA_TUNEL_1".VIBRADOR_TUNEL_1_MANUAL )
   END_RUNG
   RUNG wire#powerrail
      Contact( "BOTONERA_HMI_TUNEL_1".KM4_STOP_MANUAL_VIBRADOR_TUNEL_1 )
      wire#w1
      R_Coil( "PERMISOS_DE_MARCHA_TUNEL_1".VIBRADOR_TUNEL_1_MANUAL )
   END_RUNG
   RUNG wire#powerrail
      I_Contact( "Señal_de_fallo_vibrador_tunel_1" )
   END_RUNG wire#w1
   RUNG wire#powerrail
      Contact( "Modo_Automatico_Tunel_1" )
   END_RUNG wire#w1
   RUNG wire#powerrail
      Contact( "MEMORIAS_DE_ESTADOS_TUNEL_1".CAMBIO_ESTADO_TUNEL_1_PRESENTE )
   END_RUNG wire#w1
   RUNG wire#powerrail
      I_Contact( "Paro_Emergencia_Tunel_1" )
   END_RUNG wire#w1
   RUNG wire#powerrail
      I_Contact( "PERMISOS_GENERALES".MODO_LOCAL_1 )
   END_RUNG wire#w1
   // the same network as SCL:
   IF "BOTONERA_HMI_TUNEL_1".KM4_INICIO_MANUAL_VIBRADOR_TUNEL_1 AND "Señal_de_fallo_vibrador_tunel_1" AND "Paro_Emergencia_Tunel_1" AND "PERMISOS_GENERALES".MODO_LOCAL_1 THEN
       "PERMISOS_DE_MARCHA_TUNEL_1".VIBRADOR_TUNEL_1_MANUAL := TRUE;
   END_IF;
   IF "BOTONERA_HMI_TUNEL_1".KM4_STOP_MANUAL_VIBRADOR_TUNEL_1 OR NOT "Señal_de_fallo_vibrador_tunel_1" OR "Modo_Automatico_Tunel_1" OR "MEMORIAS_DE_ESTADOS_TUNEL_1".CAMBIO_ESTADO_TUNEL_1_PRESENTE OR NOT "Paro_Emergencia_Tunel_1" OR NOT "PERMISOS_GENERALES".MODO_LOCAL_1 THEN
       "PERMISOS_DE_MARCHA_TUNEL_1".VIBRADOR_TUNEL_1_MANUAL := FALSE;
   END_IF;
END_REGION

REGION Network 6: ABRIR CUCHARA TUNEL 1 MODO MANUAL